// TIA Portal project "ProjektZaliczenie" (V13)

(* hardware
DEVICE "HMI_1"  KTP700 Basic PN
   slot 0: "HMI"  HMI  6AV2 123-2GB03-0AX0  13.0.0.0
   slot 1: "HMI_RT_1"  KTP700 Basic PN  6AV2 123-2GB03-0AX0  13.0.0.0
   slot 5: "HMI_1.IE_CP_1"  PROFINET Interface
      slot 1: "PROFINET Interface_1"  PROFINET Interface
         slot 1: "Port_1"  Port
DEVICE "HMI_2"  KTP700 Basic PN
   slot 0: "HMI"  HMI  6AV2 123-2GB03-0AX0  13.0.1.0
   slot 1: "HMI_RT_3"  KTP700 Basic PN  6AV2 123-2GB03-0AX0  13.0.1.0
   slot 5: "HMI_2.IE_CP_1"  PROFINET Interface
      slot 1: "PROFINET Interface_1"  PROFINET Interface
         slot 1: "Port_1"  Port
DEVICE "S7-1200 station_1"  S7-1200 Station
   slot 0: "Rack_0"  Rack  V1.0
   slot 1: "PLC_1x"  CPU 1214C DC/DC/DC  6ES7 214-1AE30-0XB0  V2.2
*)

// ===== PLC "PLC_1x"  CPU 1214C DC/DC/DC =====

VAR_GLOBAL   // PLC tag table "Default tag table_1"
   "M0" AT %M1.0 : Bool;   // Zmienna pomocnicza
   "M1" AT %M1.1 : Bool;   // Zmienna pomocnicza
   "RET_VAL" AT %MW2 : Word;   // Zmienna pomocnicza
END_VAR

VAR_GLOBAL CONSTANT   // PLC tag table "Default tag table_1"
   "Local(1)" : Hw_SubModule := 50;
   "Local~PROFINET_interface_1(1)" : Hw_Interface := 64;
   "Local~PROFINET_interface_1~Port_1(1)" : Hw_Interface := 65;
   "Local~HSC_1(1)" : Hw_Hsc := 257;
   "Local~HSC_2(1)" : Hw_Hsc := 258;
   "Local~HSC_3(1)" : Hw_Hsc := 259;
   "Local~HSC_4(1)" : Hw_Hsc := 260;
   "Local~HSC_5(1)" : Hw_Hsc := 261;
   "Local~HSC_6(1)" : Hw_Hsc := 262;
   "Local~AI_2_1(1)" : Hw_SubModule := 263;
   "Local~DI_14_DQ_10_1(1)" : Hw_SubModule := 264;
   "Local~Pulse_1(1)" : Hw_Pwm := 265;
   "Local~Pulse_2(1)" : Hw_Pwm := 266;
   "OB_Main(1)" : OB_PCYCLE := 1;
   "OB_Startup(1)" : OB_STARTUP := 100;
   "RandomName" : DB_WWW := 333;
   "Local~Pulse_3" : Hw_Pwm := 267;
   "Local~Pulse_4" : Hw_Pwm := 268;
   "None" : Pip := 65535;
   "Automatic update" : Pip := 0;
   "PIP 1" : Pip := 1;
   "PIP 2" : Pip := 2;
   "PIP 3" : Pip := 3;
   "PIP 4" : Pip := 4;
   "PIP OB Servo" : Pip := 32768;
END_VAR

DATA_BLOCK "Player1DataBlock"   // DB1
{ S7_Optimized_Access := 'FALSE' }
VERSION : 0.1
   VAR
      GraphicsTypes : Array[0..99] of Int;
      EnemyBoard : Array[0..99] of Int;
      SelectedPosition : Int;
      Orientation : Bool;
      SelectedSize : Int;
      ResetAll : Bool;
      FieldsTypes : Array[0..99] of Int;
      Size4Count : Int;
      Size3Count : Int;
      Size2Count : Int;
      Size1Count : Int;
      ShipsReady : Bool;
      HP : Int;
      ReadyForNewGame : Bool;
      PlayerReady : Bool;
   END_VAR
BEGIN
END_DATA_BLOCK

DATA_BLOCK "MainDataBlock"   // DB2
{ S7_Optimized_Access := 'FALSE' }
VERSION : 0.1
   VAR
      Restart : Bool;
      JobMailBox : Array[0..3] of Word;
      Turn : Bool;
      GameResult : Int;
      JobMailBox2 : Array[0..3] of Word;
      Player1Won : Bool;
      Player2Won : Bool;
      Stage : Int;
   END_VAR
BEGIN
END_DATA_BLOCK

DATA_BLOCK "Stage1_DB"   // DB3
{ S7_Optimized_Access := 'FALSE' }
VERSION : 0.1
// stored: InstanceOfName Stage1
"Stage1"
BEGIN
END_DATA_BLOCK

DATA_BLOCK "Player2DataBlock"   // DB4
{ S7_Optimized_Access := 'FALSE' }
VERSION : 0.1
   VAR
      GraphicsTypes : Array[0..99] of Int;
      SelectedPosition : Int;
      Orientation : Bool;
      SelectedSize : Int;
      ResetAll : Bool;
      FieldsTypes : Array[0..99] of Int;
      Size4Count : Int;
      Size3Count : Int;
      Size2Count : Int;
      Size1Count : Int;
      ShipsReady : Bool;
      EnemyBoard : Array[0..99] of Int;
      HP : Int;
      ReadyForNewGame : Bool;
      PlayerReady : Bool;
   END_VAR
BEGIN
END_DATA_BLOCK

DATA_BLOCK "Stage2_DB"   // DB5
{ S7_Optimized_Access := 'FALSE' }
VERSION : 0.1
// stored: InstanceOfName Stage2
"Stage2"
BEGIN
END_DATA_BLOCK

DATA_BLOCK "Stage3_DB"   // DB6
{ S7_Optimized_Access := 'FALSE' }
VERSION : 0.1
// stored: InstanceOfName Stage3
"Stage3"
BEGIN
END_DATA_BLOCK

DATA_BLOCK "RestartGame_DB"   // DB7
{ S7_Optimized_Access := 'FALSE' }
VERSION : 0.1
// stored: InstanceOfName RestartGame
"RestartGame"
BEGIN
END_DATA_BLOCK

DATA_BLOCK "ResetShips_DB"   // DB8
{ S7_Optimized_Access := 'FALSE' }
VERSION : 0.1
// stored: InstanceOfName ResetShips
"ResetShips"
BEGIN
END_DATA_BLOCK

DATA_BLOCK "ResetShips_DB_1"   // DB9
{ S7_Optimized_Access := 'FALSE' }
VERSION : 0.1
// stored: InstanceOfName ResetShips
"ResetShips"
BEGIN
END_DATA_BLOCK

FUNCTION_BLOCK "Stage1"   // FB1, LAD
TITLE = Etap 1
{ S7_Optimized_Access := 'FALSE' }
VERSION : 0.1
// Rozmieszczanie statków przez graczy
   VAR_TEMP   // added for the SCL form of the ladder/FBD networks
      _w1 : Bool;
      _w2 : Bool;
      _w3 : Bool;
   END_VAR
BEGIN

REGION Network 1: Gracz 1
   // W momencie klniknięcia przez użytkownika na komórke (pod warunkiem wybrania rozmiaru okrętu) wywoływana jest funkcja "CheckPosition" sprawdzająca czy w wybranej lokacji można rozmieścić okręt.
   // Nastepnie, jeżeli miejsce jest dozwolone przez zasady gry, statek jest rysowany na planszy oraz inkrementowana jest aktualna ilość rozmieszczonych okrętów.
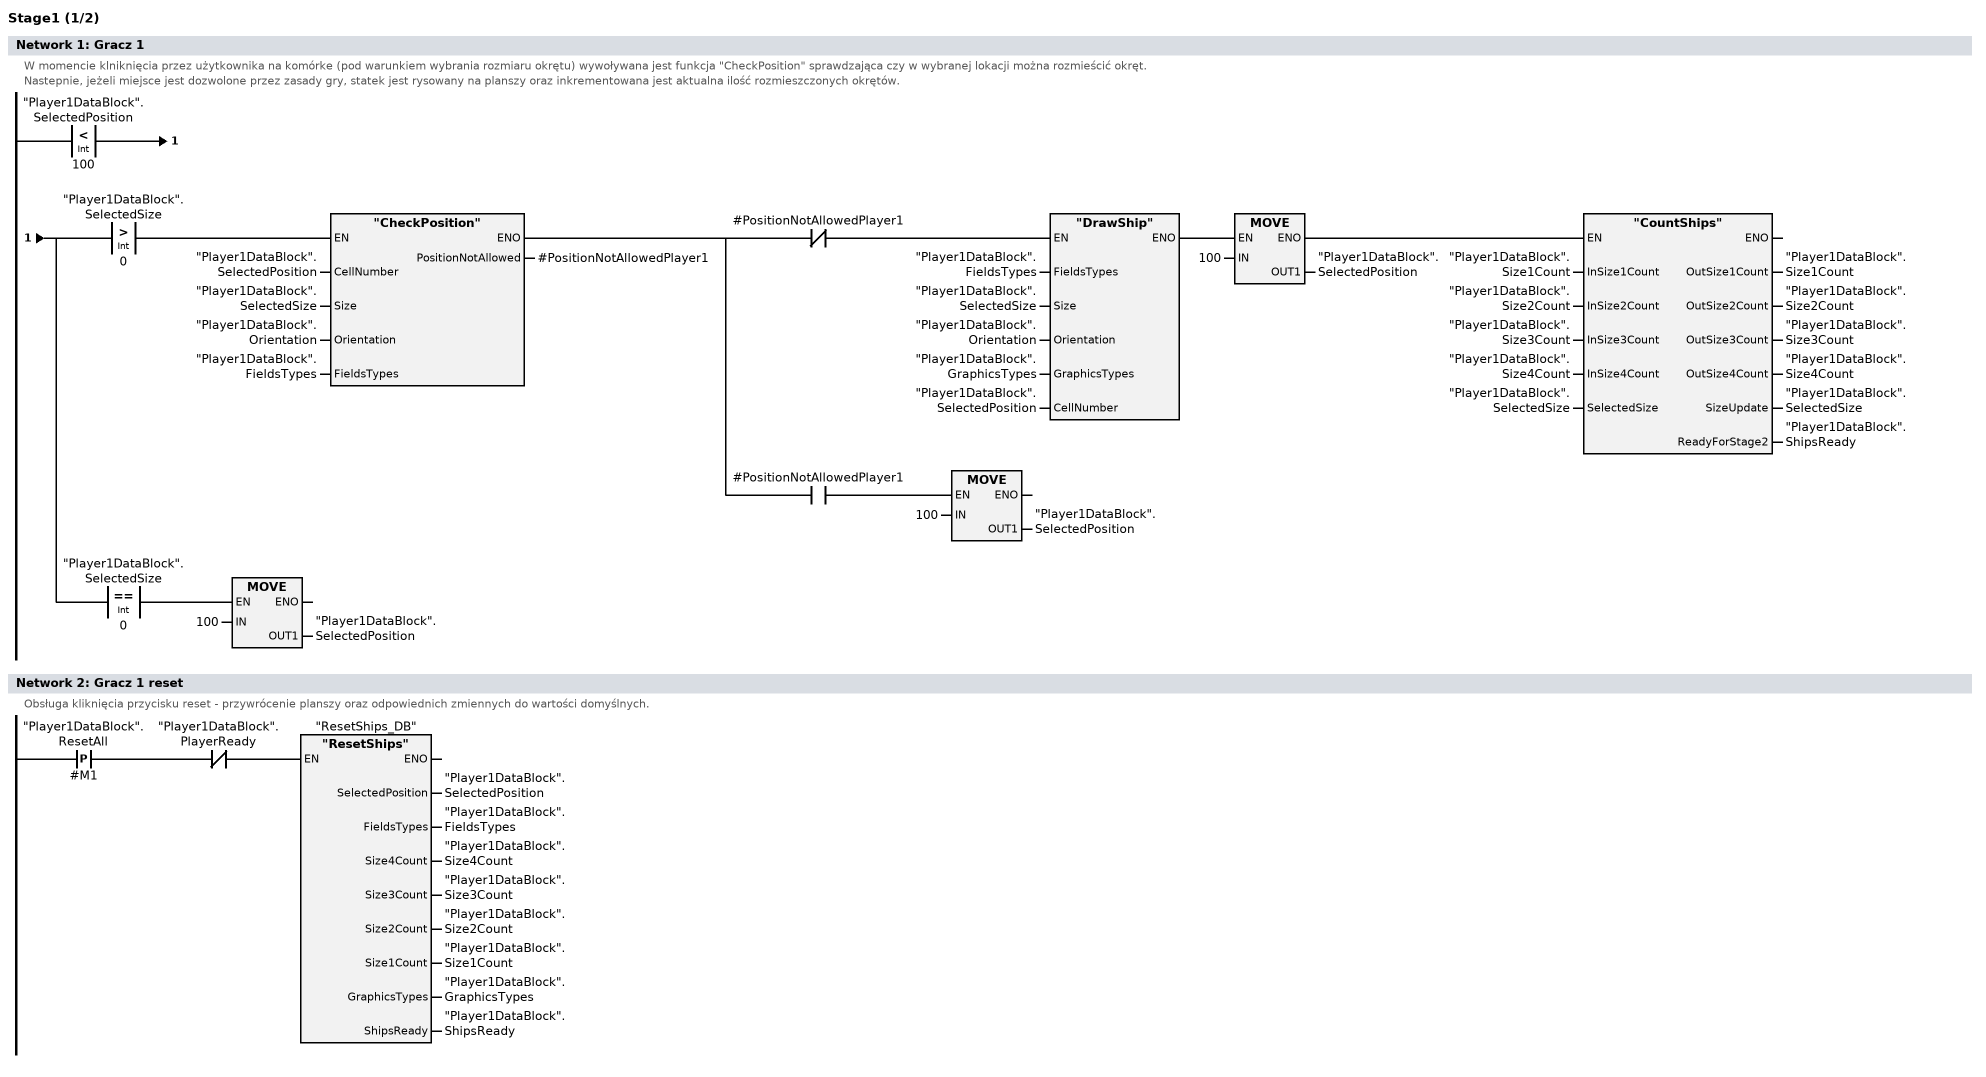
   RUNG wire#powerrail
      { S7_Templates := "SrcType := Int" } LT_Contact(in1 := "Player1DataBlock".SelectedPosition, in2 := 100)
      wire#w1
      { S7_Templates := "SrcType := Int" } GT_Contact(in1 := "Player1DataBlock".SelectedSize, in2 := 0)
      "CheckPosition"(CellNumber := "Player1DataBlock".SelectedPosition, Size := "Player1DataBlock".SelectedSize, Orientation := "Player1DataBlock".Orientation, FieldsTypes := "Player1DataBlock".FieldsTypes, PositionNotAllowed => #PositionNotAllowedPlayer1)
      wire#w2
      I_Contact( #PositionNotAllowedPlayer1 )
      "DrawShip"(FieldsTypes := "Player1DataBlock".FieldsTypes, Size := "Player1DataBlock".SelectedSize, Orientation := "Player1DataBlock".Orientation, GraphicsTypes := "Player1DataBlock".GraphicsTypes, CellNumber := "Player1DataBlock".SelectedPosition)
      Move(in := 100, out1 => "Player1DataBlock".SelectedPosition)
      "CountShips"(InSize1Count := "Player1DataBlock".Size1Count, InSize2Count := "Player1DataBlock".Size2Count, InSize3Count := "Player1DataBlock".Size3Count, InSize4Count := "Player1DataBlock".Size4Count, SelectedSize := "Player1DataBlock".SelectedSize, OutSize1Count => "Player1DataBlock".Size1Count, OutSize2Count => "Player1DataBlock".Size2Count, OutSize3Count => "Player1DataBlock".Size3Count, OutSize4Count => "Player1DataBlock".Size4Count, SizeUpdate => "Player1DataBlock".SelectedSize, ReadyForStage2 => "Player1DataBlock".ShipsReady)
   END_RUNG
   RUNG wire#w2
      Contact( #PositionNotAllowedPlayer1 )
      Move(in := 100, out1 => "Player1DataBlock".SelectedPosition)
   END_RUNG
   RUNG wire#w1
      { S7_Templates := "SrcType := Int" } EQ_Contact(in1 := "Player1DataBlock".SelectedSize, in2 := 0)
      Move(in := 100, out1 => "Player1DataBlock".SelectedPosition)
   END_RUNG
   // the same network as SCL:
   #_w1 := "Player1DataBlock".SelectedPosition < 100;
   "CheckPosition"(EN := #_w1 AND ("Player1DataBlock".SelectedSize > 0),
                   CellNumber := "Player1DataBlock".SelectedPosition,
                   Size := "Player1DataBlock".SelectedSize,
                   Orientation := "Player1DataBlock".Orientation,
                   FieldsTypes := "Player1DataBlock".FieldsTypes,
                   PositionNotAllowed => #PositionNotAllowedPlayer1,
                   ENO => #_w2);
   "DrawShip"(EN := #_w2 AND NOT #PositionNotAllowedPlayer1,
              FieldsTypes := "Player1DataBlock".FieldsTypes,
              Size := "Player1DataBlock".SelectedSize,
              Orientation := "Player1DataBlock".Orientation,
              GraphicsTypes := "Player1DataBlock".GraphicsTypes,
              CellNumber := "Player1DataBlock".SelectedPosition,
              ENO => #_w3);
   IF #_w3 THEN
       "Player1DataBlock".SelectedPosition := 100;
       "CountShips"(InSize1Count := "Player1DataBlock".Size1Count,
                    InSize2Count := "Player1DataBlock".Size2Count,
                    InSize3Count := "Player1DataBlock".Size3Count,
                    InSize4Count := "Player1DataBlock".Size4Count,
                    SelectedSize := "Player1DataBlock".SelectedSize,
                    OutSize1Count => "Player1DataBlock".Size1Count,
                    OutSize2Count => "Player1DataBlock".Size2Count,
                    OutSize3Count => "Player1DataBlock".Size3Count,
                    OutSize4Count => "Player1DataBlock".Size4Count,
                    SizeUpdate => "Player1DataBlock".SelectedSize,
                    ReadyForStage2 => "Player1DataBlock".ShipsReady);
   END_IF;
   IF #_w2 AND #PositionNotAllowedPlayer1 THEN "Player1DataBlock".SelectedPosition := 100; END_IF;
   IF #_w1 AND ("Player1DataBlock".SelectedSize = 0) THEN "Player1DataBlock".SelectedPosition := 100; END_IF;
END_REGION

REGION Network 2: Gracz 1 reset
   // Obsługa kliknięcia przycisku reset - przywrócenie planszy oraz odpowiednich zmiennych do wartości domyślnych.
   RUNG wire#powerrail
      P_Contact(operand := "Player1DataBlock".ResetAll, bit := #M1)
      I_Contact( "Player1DataBlock".PlayerReady )
      "ResetShips_DB"(SelectedPosition => "Player1DataBlock".SelectedPosition, FieldsTypes => "Player1DataBlock".FieldsTypes, Size4Count => "Player1DataBlock".Size4Count, Size3Count => "Player1DataBlock".Size3Count, Size2Count => "Player1DataBlock".Size2Count, Size1Count => "Player1DataBlock".Size1Count, GraphicsTypes => "Player1DataBlock".GraphicsTypes, ShipsReady => "Player1DataBlock".ShipsReady)
   END_RUNG
   // the same network as SCL:
   #_w1 := "Player1DataBlock".ResetAll AND NOT #M1;   // rising edge of "Player1DataBlock".ResetAll
   #M1 := "Player1DataBlock".ResetAll;
   IF #_w1 AND NOT "Player1DataBlock".PlayerReady THEN
       "ResetShips_DB"(SelectedPosition => "Player1DataBlock".SelectedPosition,   // "ResetShips"
                       FieldsTypes => "Player1DataBlock".FieldsTypes,
                       Size4Count => "Player1DataBlock".Size4Count,
                       Size3Count => "Player1DataBlock".Size3Count,
                       Size2Count => "Player1DataBlock".Size2Count,
                       Size1Count => "Player1DataBlock".Size1Count,
                       GraphicsTypes => "Player1DataBlock".GraphicsTypes,
                       ShipsReady => "Player1DataBlock".ShipsReady);
   END_IF;
END_REGION

REGION Network 3: Gracz 2
   // W momencie klniknięcia przez użytkownika na komórke (pod warunkiem wybrania rozmiaru okrętu) wywoływana jest funkcja "CheckPosition" sprawdzająca czy w wybranej lokacji można rozmieścić okręt.
   // Nastepnie, jeżeli miejsce jest dozwolone przez zasady gry, statek jest rysowany na planszy oraz inkrementowana jest aktualna ilość rozmieszczonych okrętów.
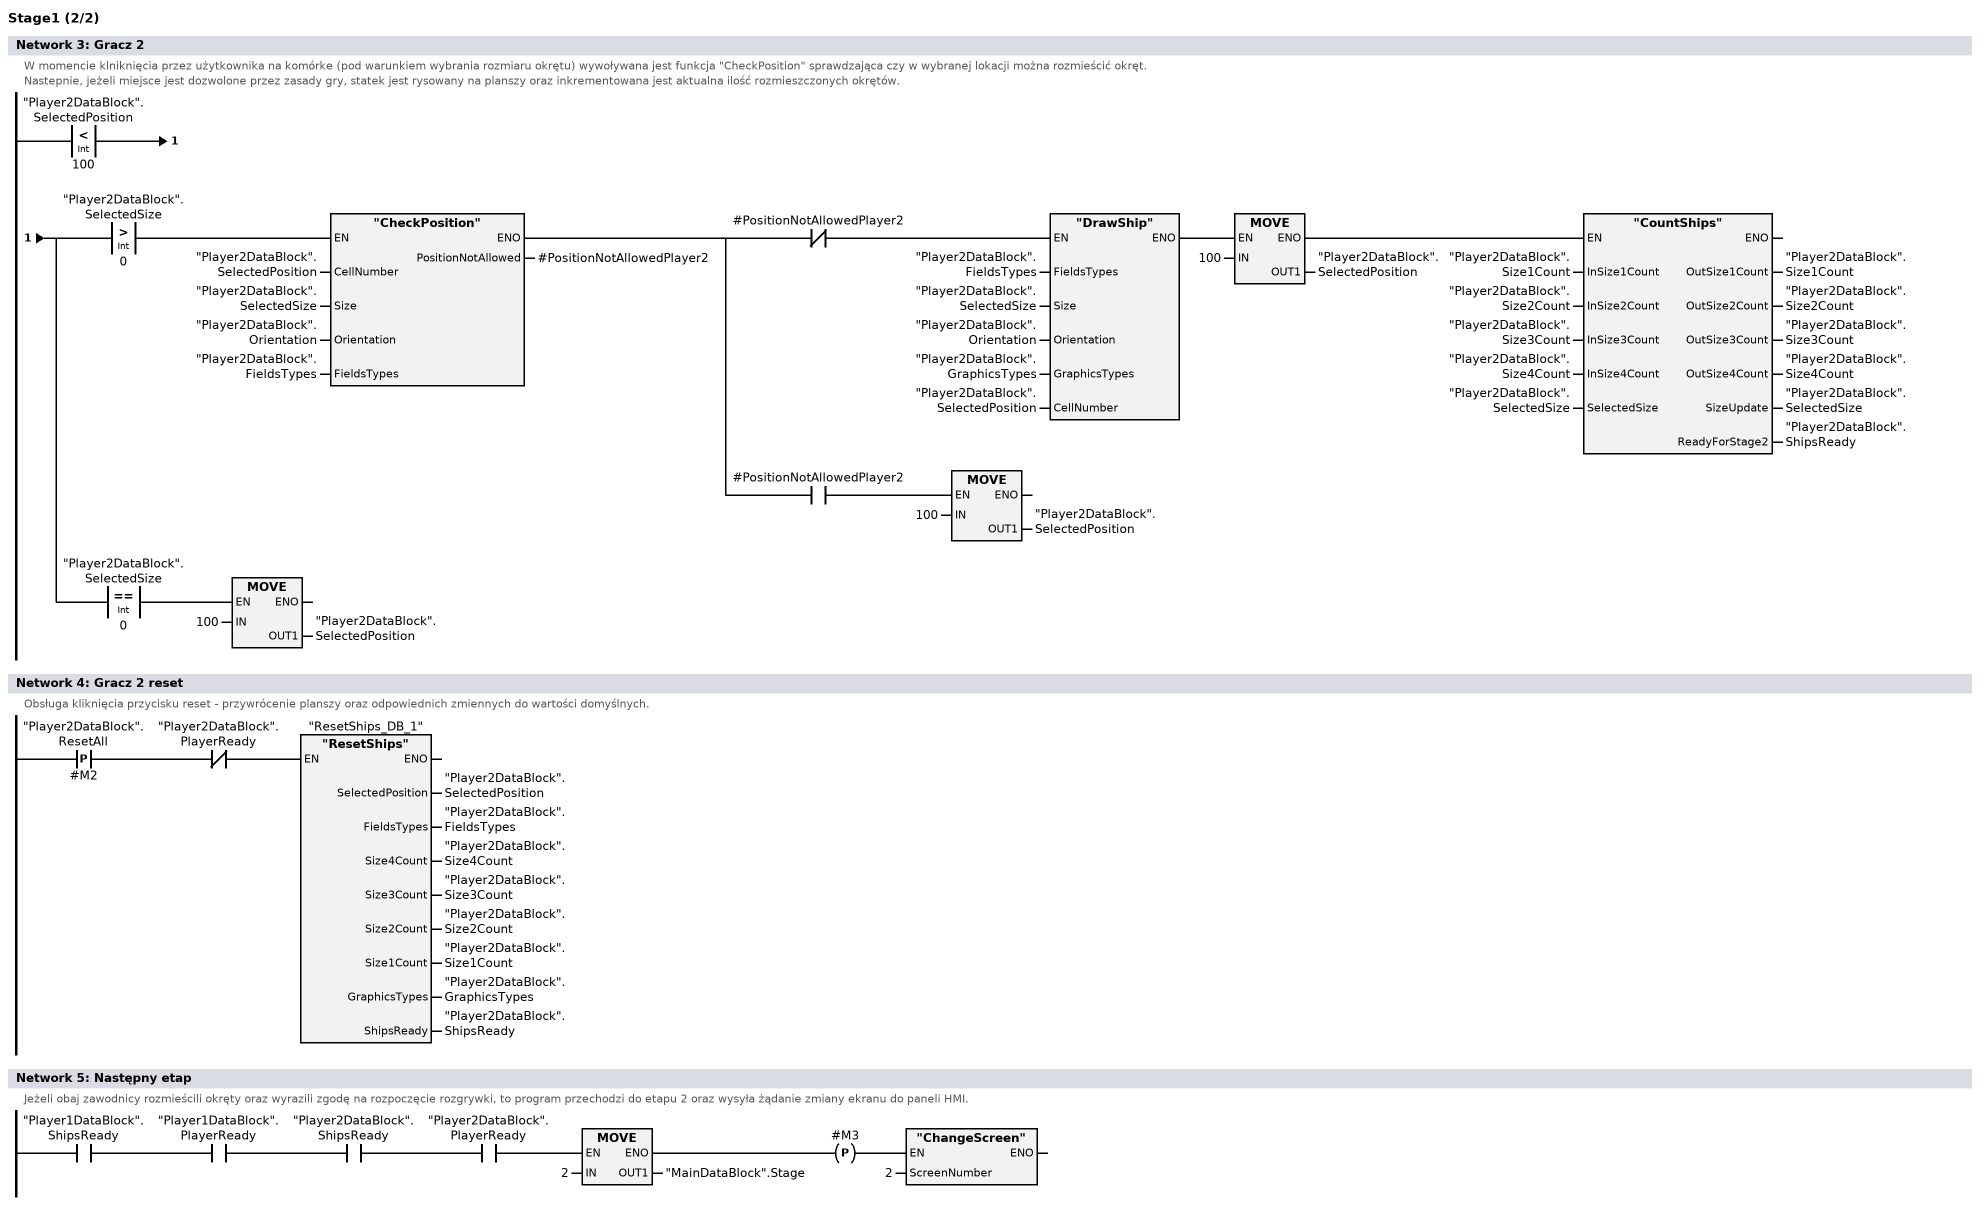
   RUNG wire#powerrail
      { S7_Templates := "SrcType := Int" } LT_Contact(in1 := "Player2DataBlock".SelectedPosition, in2 := 100)
      wire#w1
      { S7_Templates := "SrcType := Int" } GT_Contact(in1 := "Player2DataBlock".SelectedSize, in2 := 0)
      "CheckPosition"(CellNumber := "Player2DataBlock".SelectedPosition, Size := "Player2DataBlock".SelectedSize, Orientation := "Player2DataBlock".Orientation, FieldsTypes := "Player2DataBlock".FieldsTypes, PositionNotAllowed => #PositionNotAllowedPlayer2)
      wire#w2
      I_Contact( #PositionNotAllowedPlayer2 )
      "DrawShip"(FieldsTypes := "Player2DataBlock".FieldsTypes, Size := "Player2DataBlock".SelectedSize, Orientation := "Player2DataBlock".Orientation, GraphicsTypes := "Player2DataBlock".GraphicsTypes, CellNumber := "Player2DataBlock".SelectedPosition)
      Move(in := 100, out1 => "Player2DataBlock".SelectedPosition)
      "CountShips"(InSize1Count := "Player2DataBlock".Size1Count, InSize2Count := "Player2DataBlock".Size2Count, InSize3Count := "Player2DataBlock".Size3Count, InSize4Count := "Player2DataBlock".Size4Count, SelectedSize := "Player2DataBlock".SelectedSize, OutSize1Count => "Player2DataBlock".Size1Count, OutSize2Count => "Player2DataBlock".Size2Count, OutSize3Count => "Player2DataBlock".Size3Count, OutSize4Count => "Player2DataBlock".Size4Count, SizeUpdate => "Player2DataBlock".SelectedSize, ReadyForStage2 => "Player2DataBlock".ShipsReady)
   END_RUNG
   RUNG wire#w2
      Contact( #PositionNotAllowedPlayer2 )
      Move(in := 100, out1 => "Player2DataBlock".SelectedPosition)
   END_RUNG
   RUNG wire#w1
      { S7_Templates := "SrcType := Int" } EQ_Contact(in1 := "Player2DataBlock".SelectedSize, in2 := 0)
      Move(in := 100, out1 => "Player2DataBlock".SelectedPosition)
   END_RUNG
   // the same network as SCL:
   #_w1 := "Player2DataBlock".SelectedPosition < 100;
   "CheckPosition"(EN := #_w1 AND ("Player2DataBlock".SelectedSize > 0),
                   CellNumber := "Player2DataBlock".SelectedPosition,
                   Size := "Player2DataBlock".SelectedSize,
                   Orientation := "Player2DataBlock".Orientation,
                   FieldsTypes := "Player2DataBlock".FieldsTypes,
                   PositionNotAllowed => #PositionNotAllowedPlayer2,
                   ENO => #_w2);
   "DrawShip"(EN := #_w2 AND NOT #PositionNotAllowedPlayer2,
              FieldsTypes := "Player2DataBlock".FieldsTypes,
              Size := "Player2DataBlock".SelectedSize,
              Orientation := "Player2DataBlock".Orientation,
              GraphicsTypes := "Player2DataBlock".GraphicsTypes,
              CellNumber := "Player2DataBlock".SelectedPosition,
              ENO => #_w3);
   IF #_w3 THEN
       "Player2DataBlock".SelectedPosition := 100;
       "CountShips"(InSize1Count := "Player2DataBlock".Size1Count,
                    InSize2Count := "Player2DataBlock".Size2Count,
                    InSize3Count := "Player2DataBlock".Size3Count,
                    InSize4Count := "Player2DataBlock".Size4Count,
                    SelectedSize := "Player2DataBlock".SelectedSize,
                    OutSize1Count => "Player2DataBlock".Size1Count,
                    OutSize2Count => "Player2DataBlock".Size2Count,
                    OutSize3Count => "Player2DataBlock".Size3Count,
                    OutSize4Count => "Player2DataBlock".Size4Count,
                    SizeUpdate => "Player2DataBlock".SelectedSize,
                    ReadyForStage2 => "Player2DataBlock".ShipsReady);
   END_IF;
   IF #_w2 AND #PositionNotAllowedPlayer2 THEN "Player2DataBlock".SelectedPosition := 100; END_IF;
   IF #_w1 AND ("Player2DataBlock".SelectedSize = 0) THEN "Player2DataBlock".SelectedPosition := 100; END_IF;
END_REGION

REGION Network 4: Gracz 2 reset
   // Obsługa kliknięcia przycisku reset - przywrócenie planszy oraz odpowiednich zmiennych do wartości domyślnych.
   RUNG wire#powerrail
      P_Contact(operand := "Player2DataBlock".ResetAll, bit := #M2)
      I_Contact( "Player2DataBlock".PlayerReady )
      "ResetShips_DB_1"(SelectedPosition => "Player2DataBlock".SelectedPosition, FieldsTypes => "Player2DataBlock".FieldsTypes, Size4Count => "Player2DataBlock".Size4Count, Size3Count => "Player2DataBlock".Size3Count, Size2Count => "Player2DataBlock".Size2Count, Size1Count => "Player2DataBlock".Size1Count, GraphicsTypes => "Player2DataBlock".GraphicsTypes, ShipsReady => "Player2DataBlock".ShipsReady)
   END_RUNG
   // the same network as SCL:
   #_w1 := "Player2DataBlock".ResetAll AND NOT #M2;   // rising edge of "Player2DataBlock".ResetAll
   #M2 := "Player2DataBlock".ResetAll;
   IF #_w1 AND NOT "Player2DataBlock".PlayerReady THEN
       "ResetShips_DB_1"(SelectedPosition => "Player2DataBlock".SelectedPosition,   // "ResetShips"
                         FieldsTypes => "Player2DataBlock".FieldsTypes,
                         Size4Count => "Player2DataBlock".Size4Count,
                         Size3Count => "Player2DataBlock".Size3Count,
                         Size2Count => "Player2DataBlock".Size2Count,
                         Size1Count => "Player2DataBlock".Size1Count,
                         GraphicsTypes => "Player2DataBlock".GraphicsTypes,
                         ShipsReady => "Player2DataBlock".ShipsReady);
   END_IF;
END_REGION

REGION Network 5: Następny etap
   // Jeżeli obaj zawodnicy rozmieścili okręty oraz wyrazili zgodę na rozpoczęcie rozgrywki, to program przechodzi do etapu 2 oraz wysyła żądanie zmiany ekranu do paneli HMI.
   RUNG wire#powerrail
      Contact( "Player1DataBlock".ShipsReady )
      Contact( "Player1DataBlock".PlayerReady )
      Contact( "Player2DataBlock".ShipsReady )
      Contact( "Player2DataBlock".PlayerReady )
      { S7_GenerateENO := "TRUE" } Move(in := 2, out1 => "MainDataBlock".Stage)
      P_Trig( #M3 )
      "ChangeScreen"(ScreenNumber := 2)
   END_RUNG
   // the same network as SCL:
   // ENO of a box is taken as its EN; it also drops when the box reports an error
   #_w1 := "Player1DataBlock".ShipsReady AND "Player1DataBlock".PlayerReady AND "Player2DataBlock".ShipsReady AND "Player2DataBlock".PlayerReady;
   IF #_w1 THEN "MainDataBlock".Stage := 2; END_IF;
   #_w2 := #_w1 AND NOT #M3;   // rising edge
   #M3 := #_w1;
   IF #_w2 THEN "ChangeScreen"(ScreenNumber := 2); END_IF;
END_REGION
END_FUNCTION_BLOCK

FUNCTION_BLOCK "Stage2"   // FB2, LAD
TITLE = Etap 2
{ S7_Optimized_Access := 'FALSE' }
VERSION : 0.1
// Właściwa rozgrywka
   VAR_TEMP   // added for the SCL form of the ladder/FBD networks
      _w1 : Bool;
      _w2 : Bool;
      _w3 : Bool;
   END_VAR
BEGIN

REGION Network 1: Ruch gracza 1
   // Jeżeli tura należy do gracza oraz wybrał on komórkę na planszy, to sprawdzane jest trafienie poprzez funkcję "CheckHit". 
   // W przypadku trafienia gracz zyskuje możliwość ponowngeo strzału, a przeciwnikowi odejmowany jest punkt HP.
   // W przypadku pudła gracz oddaje ruch przeciwnikowi.
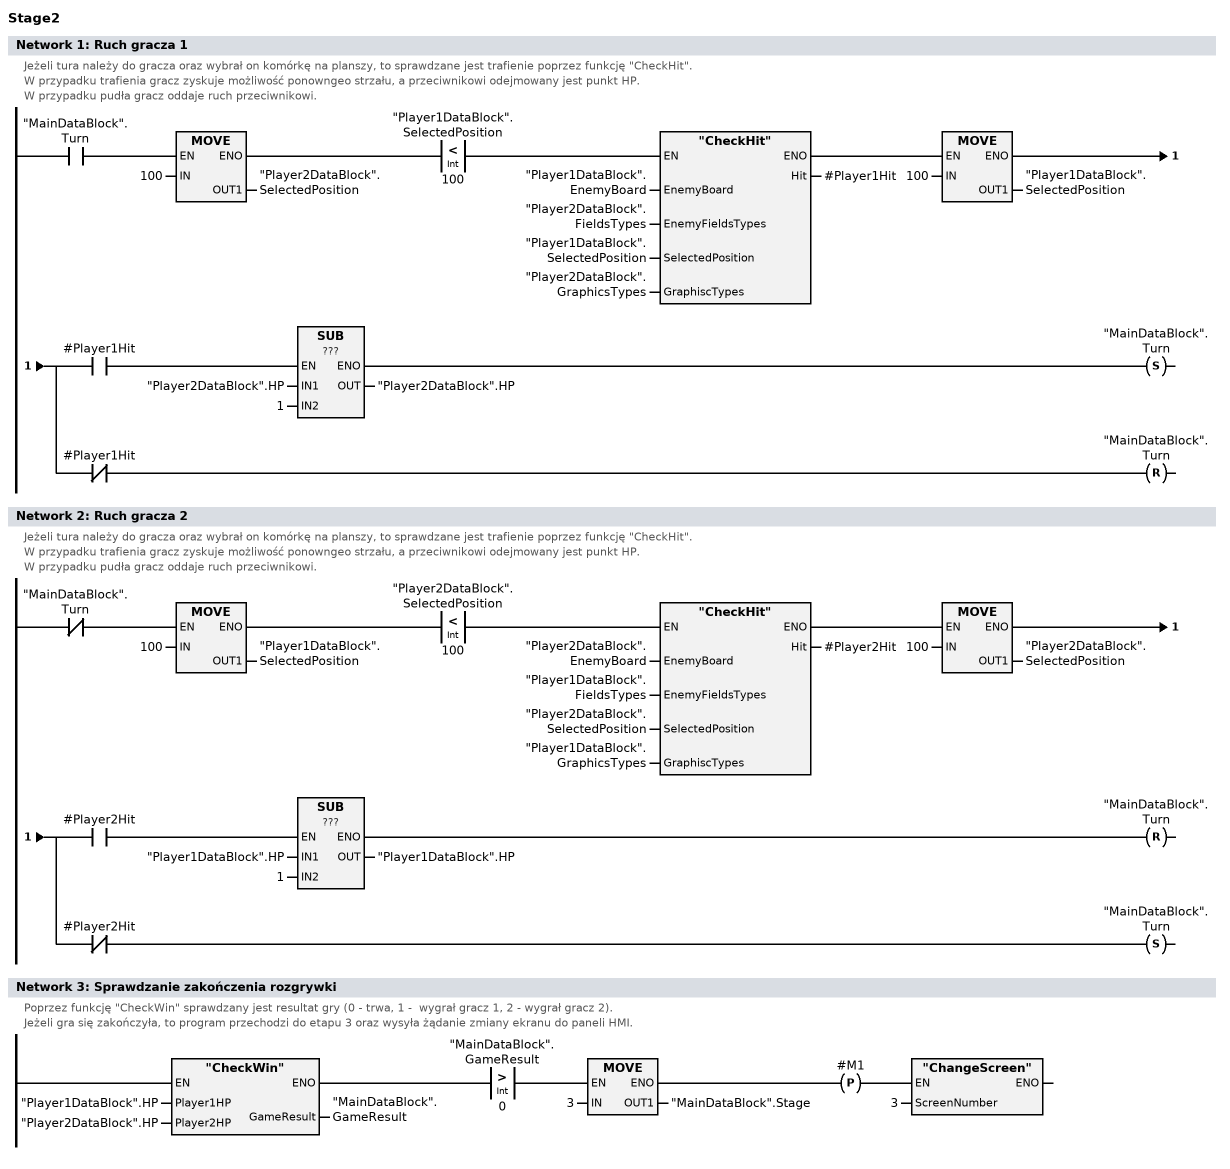
   RUNG wire#powerrail
      Contact( "MainDataBlock".Turn )
      { S7_GenerateENO := "TRUE" } Move(in := 100, out1 => "Player2DataBlock".SelectedPosition)
      { S7_Templates := "SrcType := Int" } LT_Contact(in1 := "Player1DataBlock".SelectedPosition, in2 := 100)
      "CheckHit"(EnemyBoard := "Player1DataBlock".EnemyBoard, EnemyFieldsTypes := "Player2DataBlock".FieldsTypes, SelectedPosition := "Player1DataBlock".SelectedPosition, GraphiscTypes := "Player2DataBlock".GraphicsTypes, Hit => #Player1Hit)
      { S7_GenerateENO := "TRUE" } Move(in := 100, out1 => "Player1DataBlock".SelectedPosition)
      wire#w1
      Contact( #Player1Hit )
      { S7_Templates := "SrcType := ???"; S7_GenerateENO := "TRUE" } Sub(in1 := "Player2DataBlock".HP, in2 := 1, out => "Player2DataBlock".HP)
      S_Coil( "MainDataBlock".Turn )
   END_RUNG
   RUNG wire#w1
      I_Contact( #Player1Hit )
      R_Coil( "MainDataBlock".Turn )
   END_RUNG
   // the same network as SCL:
   // ENO of a box is taken as its EN; it also drops when the box reports an error
   IF "MainDataBlock".Turn THEN "Player2DataBlock".SelectedPosition := 100; END_IF;
   "CheckHit"(EN := "MainDataBlock".Turn AND ("Player1DataBlock".SelectedPosition < 100),
              EnemyBoard := "Player1DataBlock".EnemyBoard,
              EnemyFieldsTypes := "Player2DataBlock".FieldsTypes,
              SelectedPosition := "Player1DataBlock".SelectedPosition,
              GraphiscTypes := "Player2DataBlock".GraphicsTypes,
              Hit => #Player1Hit,
              ENO => #_w1);
   IF #_w1 THEN "Player1DataBlock".SelectedPosition := 100; END_IF;
   IF #_w1 AND #Player1Hit THEN
       "Player2DataBlock".HP := "Player2DataBlock".HP - 1;
       "MainDataBlock".Turn := TRUE;
   END_IF;
   IF #_w1 AND NOT #Player1Hit THEN "MainDataBlock".Turn := FALSE; END_IF;
END_REGION

REGION Network 2: Ruch gracza 2
   // Jeżeli tura należy do gracza oraz wybrał on komórkę na planszy, to sprawdzane jest trafienie poprzez funkcję "CheckHit". 
   // W przypadku trafienia gracz zyskuje możliwość ponowngeo strzału, a przeciwnikowi odejmowany jest punkt HP.
   // W przypadku pudła gracz oddaje ruch przeciwnikowi.
   RUNG wire#powerrail
      I_Contact( "MainDataBlock".Turn )
      { S7_GenerateENO := "TRUE" } Move(in := 100, out1 => "Player1DataBlock".SelectedPosition)
      { S7_Templates := "SrcType := Int" } LT_Contact(in1 := "Player2DataBlock".SelectedPosition, in2 := 100)
      "CheckHit"(EnemyBoard := "Player2DataBlock".EnemyBoard, EnemyFieldsTypes := "Player1DataBlock".FieldsTypes, SelectedPosition := "Player2DataBlock".SelectedPosition, GraphiscTypes := "Player1DataBlock".GraphicsTypes, Hit => #Player2Hit)
      { S7_GenerateENO := "TRUE" } Move(in := 100, out1 => "Player2DataBlock".SelectedPosition)
      wire#w1
      Contact( #Player2Hit )
      { S7_Templates := "SrcType := ???"; S7_GenerateENO := "TRUE" } Sub(in1 := "Player1DataBlock".HP, in2 := 1, out => "Player1DataBlock".HP)
      R_Coil( "MainDataBlock".Turn )
   END_RUNG
   RUNG wire#w1
      I_Contact( #Player2Hit )
      S_Coil( "MainDataBlock".Turn )
   END_RUNG
   // the same network as SCL:
   // ENO of a box is taken as its EN; it also drops when the box reports an error
   IF NOT "MainDataBlock".Turn THEN "Player1DataBlock".SelectedPosition := 100; END_IF;
   "CheckHit"(EN := NOT "MainDataBlock".Turn AND ("Player2DataBlock".SelectedPosition < 100),
              EnemyBoard := "Player2DataBlock".EnemyBoard,
              EnemyFieldsTypes := "Player1DataBlock".FieldsTypes,
              SelectedPosition := "Player2DataBlock".SelectedPosition,
              GraphiscTypes := "Player1DataBlock".GraphicsTypes,
              Hit => #Player2Hit,
              ENO => #_w1);
   IF #_w1 THEN "Player2DataBlock".SelectedPosition := 100; END_IF;
   IF #_w1 AND #Player2Hit THEN
       "Player1DataBlock".HP := "Player1DataBlock".HP - 1;
       "MainDataBlock".Turn := FALSE;
   END_IF;
   IF #_w1 AND NOT #Player2Hit THEN "MainDataBlock".Turn := TRUE; END_IF;
END_REGION

REGION Network 3: Sprawdzanie zakończenia rozgrywki
   // Poprzez funkcję "CheckWin" sprawdzany jest resultat gry (0 - trwa, 1 -  wygrał gracz 1, 2 - wygrał gracz 2). 
   // Jeżeli gra się zakończyła, to program przechodzi do etapu 3 oraz wysyła żądanie zmiany ekranu do paneli HMI.
   RUNG wire#powerrail
      "CheckWin"(Player1HP := "Player1DataBlock".HP, Player2HP := "Player2DataBlock".HP, GameResult => "MainDataBlock".GameResult)
      { S7_Templates := "SrcType := Int" } GT_Contact(in1 := "MainDataBlock".GameResult, in2 := 0)
      { S7_GenerateENO := "TRUE" } Move(in := 3, out1 => "MainDataBlock".Stage)
      P_Trig( #M1 )
      "ChangeScreen"(ScreenNumber := 3)
   END_RUNG
   // the same network as SCL:
   // ENO of a box is taken as its EN; it also drops when the box reports an error
   "CheckWin"(Player1HP := "Player1DataBlock".HP,
              Player2HP := "Player2DataBlock".HP,
              GameResult => "MainDataBlock".GameResult,
              ENO => #_w1);
   #_w2 := #_w1 AND ("MainDataBlock".GameResult > 0);
   IF #_w2 THEN "MainDataBlock".Stage := 3; END_IF;
   #_w3 := #_w2 AND NOT #M1;   // rising edge
   #M1 := #_w2;
   IF #_w3 THEN "ChangeScreen"(ScreenNumber := 3); END_IF;
END_REGION
END_FUNCTION_BLOCK

FUNCTION_BLOCK "Stage3"   // FB3, LAD
TITLE = Etap 3
{ S7_Optimized_Access := 'FALSE' }
VERSION : 0.1
// Wyświetlenie wyniku starcia oraz oczekiwanie na nawą rozgrywkę.
   VAR_TEMP   // added for the SCL form of the ladder/FBD networks
      _w1 : Bool;
      _w2 : Bool;
   END_VAR
BEGIN

REGION Network 1: Sprawdzanie czy gracze są gotowi na nową rozgrywkę
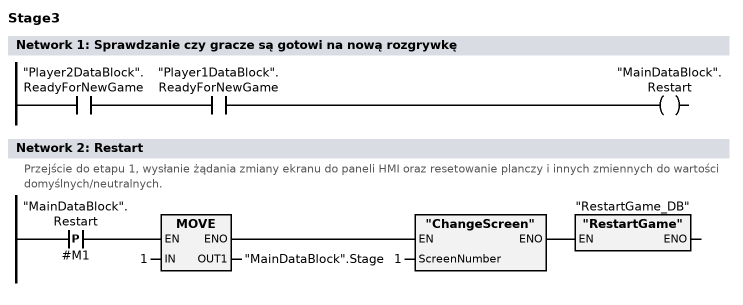
   RUNG wire#powerrail
      Contact( "Player2DataBlock".ReadyForNewGame )
      Contact( "Player1DataBlock".ReadyForNewGame )
      Coil( "MainDataBlock".Restart )
   END_RUNG
   // the same network as SCL:
   "MainDataBlock".Restart := "Player2DataBlock".ReadyForNewGame AND "Player1DataBlock".ReadyForNewGame;
END_REGION

REGION Network 2: Restart
   // Przejście do etapu 1, wysłanie żądania zmiany ekranu do paneli HMI oraz resetowanie planczy i innych zmiennych do wartości domyślnych/neutralnych.
   RUNG wire#powerrail
      P_Contact(operand := "MainDataBlock".Restart, bit := #M1)
      { S7_GenerateENO := "TRUE" } Move(in := 1, out1 => "MainDataBlock".Stage)
      "ChangeScreen"(ScreenNumber := 1)
      "RestartGame_DB"()
   END_RUNG
   // the same network as SCL:
   // ENO of a box is taken as its EN; it also drops when the box reports an error
   #_w1 := "MainDataBlock".Restart AND NOT #M1;   // rising edge of "MainDataBlock".Restart
   #M1 := "MainDataBlock".Restart;
   IF #_w1 THEN "MainDataBlock".Stage := 1; END_IF;
   "ChangeScreen"(EN := #_w1, ScreenNumber := 1, ENO => #_w2);
   IF #_w2 THEN
       "RestartGame_DB"();   // "RestartGame"
   END_IF;
END_REGION
END_FUNCTION_BLOCK

FUNCTION_BLOCK "RestartGame"   // FB4, LAD
TITLE = Restartowanie rozgrywki
{ S7_Optimized_Access := 'FALSE' }
VERSION : 0.1
BEGIN

REGION Network 1: Resetowanie wartości zmiennych (ustawianie wartości domyślnych/neutralnych)